                           REGION "RED OFF"
                               IF NOT "Clock_1Hz" THEN
                                   CASE #j OF
                                       #"Part 01":
                                           #stackLight := #stackLight AND (NOT #"Part 01 Red On");
                                           #stackLight := #stackLight AND (NOT #"Part 01 Yellow On");
                                           #stackLight := #stackLight AND (NOT #"Part 01 Green On");
                                       #"Part 02":
                                           #stackLight := #stackLight AND (NOT #"Part 02 Red On");
                                           #stackLight := #stackLight AND (NOT #"Part 02 Yellow On");
                                           #stackLight := #stackLight AND (NOT #"Part 02 Green On");
                                       #"Part 03":
                                           #stackLight := #stackLight AND (NOT #"Part 03 Red On");
                                           #stackLight := #stackLight AND (NOT #"Part 03 Yellow On");
                                           #stackLight := #stackLight AND (NOT #"Part 03 Green On");
                                       #"Part 04":
                                           #stackLight := #stackLight AND (NOT #"Part 04 Red On");
                                           #stackLight := #stackLight AND (NOT #"Part 04 Yellow On");
                                           #stackLight := #stackLight AND (NOT #"Part 04 Green On");
                                       #"Part 05":
                                           #stackLight := #stackLight AND (NOT #"Part 05 Red On");
                                           #stackLight := #stackLight AND (NOT #"Part 05 Yellow On");
                                           #stackLight := #stackLight AND (NOT #"Part 05 Green On");
                                       #"Part 06":
                                           #stackLight := #stackLight AND (NOT #"Part 06 Red On");
                                           #stackLight := #stackLight AND (NOT #"Part 06 Yellow On");
                                           #stackLight := #stackLight AND (NOT #"Part 06 Green On");
                                       ELSE
                                           ;
                                   END_CASE;
                               END_IF;
                           END_REGION

                       END_IF;
                   END_REGION

                   REGION "COPY OUT TO GLOBAL"
                       #stations.me[#i].stackLightOut := #stackLight;
                   END_REGION

               END_FOR;
           END_REGION

       END_FOR;
   END_REGION
END_FUNCTION_BLOCK

FUNCTION_BLOCK "KP8 Button Activation"   // FB12, SCL
{ S7_Optimized_Access := 'TRUE' }
VERSION : 0.1
   VAR_IN_OUT
      stations : "Stations";
   END_VAR
   VAR
      old : Struct
         kp8Config : Array[0.."stnCount"] of "KP8 Button Config";
      END_STRUCT;
   END_VAR
   VAR_TEMP
      btnCount : Int;
      currentPNs : Array[0..7] of WString[40];
      i : Int;
      init : Bool;
      j : Int;
      stnCount : Int;
      temp : Int;
   END_VAR
BEGIN
   REGION "GET STATION COUNT"
       #stnCount := "stnCount";
       #btnCount := "ptsPerStn";
   END_REGION

   REGION "LOOP THROUGH STATIONS"
       FOR #i := 0 TO #stnCount DO

           REGION "COPY TO LOCAL"
               #currentPNs := #stations.me[#i].partNumbers;
           END_REGION


           REGION "LOOP THROUGH BUTTONS"
               FOR #j := 0 TO #btnCount DO

                       REGION "ACTIVATE BUTTON"
                           IF LEN(#currentPNs[#j]) <> 0 THEN
                               #stations.me[#i].kp8Config.activate[#j] := TRUE;
                               #stations.me[#i].kp8Config.colorOff[#j] := 'green';
                               #stations.me[#i].kp8Config.colorOn1[#j] := 'yellow';
                               #stations.me[#i].kp8Config.colorOn2[#j] := '';
                               #stations.me[#i].kp8Config.flash[#j] := FALSE;
                               #stations.me[#i].kp8Config.group[#j] := 0;
                               #stations.me[#i].kp8Config.mode[#j] := TRUE;
                           END_IF;
                       END_REGION

                       REGION "DEACTIVATE BUTTON"
                           IF LEN(#currentPNs[#j]) = 0 THEN
                               #stations.me[#i].kp8Config.activate[#j] := FALSE;
                               #stations.me[#i].kp8Config.colorOff[#j] := '';
                               #stations.me[#i].kp8Config.colorOn1[#j] := '';
                               #stations.me[#i].kp8Config.colorOn2[#j] := '';
                               #stations.me[#i].kp8Config.flash[#j] := FALSE;
                               #stations.me[#i].kp8Config.group[#j] := 0;
                               #stations.me[#i].kp8Config.mode[#j] := FALSE;
                           END_IF;
                       END_REGION

               END_FOR;
           END_REGION

           REGION "SOFT INIT"
               IF #stations.me[#i].kp8Config <> #old.kp8Config[#i] THEN
                   #stations.me[#i].init.soft := TRUE;
               END_IF;
           END_REGION

           REGION "SAVE FOR CHANGE DETECTION"
               #old.kp8Config[#i] := #stations.me[#i].kp8Config;
           END_REGION

       END_FOR;
   END_REGION
END_FUNCTION_BLOCK

FUNCTION_BLOCK "Remove Part Request"   // FB13, SCL
{ S7_Optimized_Access := 'TRUE' }
VERSION : 0.1
   VAR_IN_OUT
      pRow : Int;
      requests : "Part Request Data";
      stations : "Stations";
   END_VAR
   VAR
      old : Struct
         partReq : "Station Old Presses";
      END_STRUCT;
   END_VAR
   VAR_TEMP
      address : UInt;
      blankRow : "Table Row";
      hasPart : Bool;
      i : Int;
      j : Int;
      k : Int;
      logAddress : UInt;
      maxRows : Int;
      noPart : Bool;
      oldPartReq : Bool;
      partNumber : WString;
      partReq : Bool;
      pRemoveRow : Int;
      btnCount : Int;
      stnCount : Int;
      removeAddress : Bool;
   END_VAR
BEGIN
   REGION "COPY TO LOCAL"
       #maxRows := "partReqHmiRowCount";
       #stnCount := "stnCount";
       #btnCount := "ptsPerStn";
   END_REGION


   REGION "FOR EACH STATION"
       FOR #i := 0 TO #stnCount DO

           REGION "FOR EACH BUTTON"
               FOR #j := 1 TO #btnCount DO

                   REGION "COPY TO LOCAL"
                       #partReq := #stations.me[#i].btnStates[#j];
                       #oldPartReq := #old.partReq.me[#i, #j];
                   END_REGION

                   REGION "DETERMINE STATE"

                       REGION "PART REQUEST FALLING EDGE"
                           IF NOT #partReq AND #oldPartReq THEN

                               REGION "SAVE FOR CHANGE DETECTION"
                                   #old.partReq.me[#i, #j] := #partReq;
                               END_REGION

                               REGION "COPY TO LOCAL"
                                   #partNumber := #stations.me[#i].partNumbers[#j];
                               END_REGION

                               REGION "BUTTON HAS NO PART"
                                   IF #partNumber = wstring#'' THEN
                                       #hasPart := FALSE;
                                       #noPart := TRUE;
                                   END_IF;
                               END_REGION

                               REGION "BUTTON HAS PART"
                                   IF #partNumber <> wstring#'' THEN
                                       #hasPart := TRUE;
                                       #noPart := FALSE;
                                   END_IF;
                               END_REGION

                           END_IF;
                       END_REGION

                   END_REGION

                   REGION "NO PART"
                       IF #noPart THEN

                           REGION "TURN OFF THE LIGHTS"
                               #hasPart := FALSE;
                               #noPart := FALSE;
                           END_REGION

                       END_IF;

                   END_REGION

                   REGION "HAS PART"
                       IF #hasPart THEN

                           REGION "TURN OFF THE LIGHTS"
                               #hasPart := FALSE;
                           END_REGION

                           REGION "CALCULATE ADDRESS"
                               #address := (INT_TO_UINT(#i) + 1) * 10 + (INT_TO_UINT(#j) + 1);
                           END_REGION

                           REGION "RESET FLAG"
                               #removeAddress := FALSE;
                           END_REGION

                           REGION "SEARCH EACH ROW IN PART DB"
                               FOR #k := 0 TO #maxRows DO

                                   REGION "COPY TO LOCAL"
                                       #logAddress := #requests.row[#k].address;
                                   END_REGION

                                   REGION "ON MATCH"
                                       IF #logAddress = #address THEN

                                           REGION "SET FLAG"
                                               #removeAddress := TRUE;
                                           END_REGION

                                           REGION "SAVE POINTER"
                                               #pRemoveRow := #k;
                                           END_REGION

                                       END_IF;
                                   END_REGION

                               END_FOR;
                           END_REGION

                       END_IF;
                   END_REGION

                   REGION "REMOVE ADDRESS"
                       IF #removeAddress THEN

                           REGION "TURN OFF THE LIGHTS"
                               #removeAddress := FALSE;
                           END_REGION

                           REGION "TURN OFF REQUEST"
                               #stations.me[#i].partRequested[#j] := FALSE;
                           END_REGION

                           REGION "REMOVAL PROCESS"

                               REGION "REMOVE ROW"
                                   #requests.row[#pRemoveRow] := #blankRow;
                               END_REGION

                               REGION "REMOVE PART ORDERED"
                                   #stations.me[#i].partOrdered[#j] := FALSE;
                               END_REGION

                           END_REGION

                           REGION "ROW POINTER"

                               REGION "DECREMENT"
                                   #pRow := #pRow - 1;
                               END_REGION

                               REGION "LOW LIMIT ROLL OVER"
                                   IF #pRow < 0 THEN
                                       #pRow := 0;
                                   END_IF;
                               END_REGION

                           END_REGION

                       END_IF;
                   END_REGION

               END_FOR;

           END_REGION

       END_FOR;
   END_REGION
END_FUNCTION_BLOCK

FUNCTION_BLOCK "HMI Settings Screen"   // FB14, LAD
{ S7_Optimized_Access := 'TRUE' }
VERSION : 0.1
   VAR_IN_OUT
      settings : "Settings";
      stations : "Stations";
   END_VAR
   VAR
      tmrTimeOut : TON_TIME;
      instStaSel : "Station Selection";
      instKP8BtnSel : "KP8 Button Selections";
      old : Struct
         asgnPN : Bool;
         asgnAlloted : Bool;
         asgnCritical : Bool;
         nextPress : Bool;
         prevPress : Bool;
         selBtnCount : Int;
         selBtnNumber : Int;
         selStnCount : Int;
         selStnNumber : Int;
      END_STRUCT;
      instAsnBtnPrms : "Assign Button Parameters";
      instAniPNTmr : "Animate: PN & Timers";
   END_VAR
   VAR_TEMP
      pBN : Int;
      pSN : Int;
      wStringBox : WString;
   END_VAR
   VAR CONSTANT
      ptTimeOut : Time := t#15m;
   END_VAR
   VAR_TEMP   // added for the SCL form of the ladder/FBD networks
      _w1 : Bool;
   END_VAR
BEGIN

REGION Network 1: ENTRY TIMEOUT
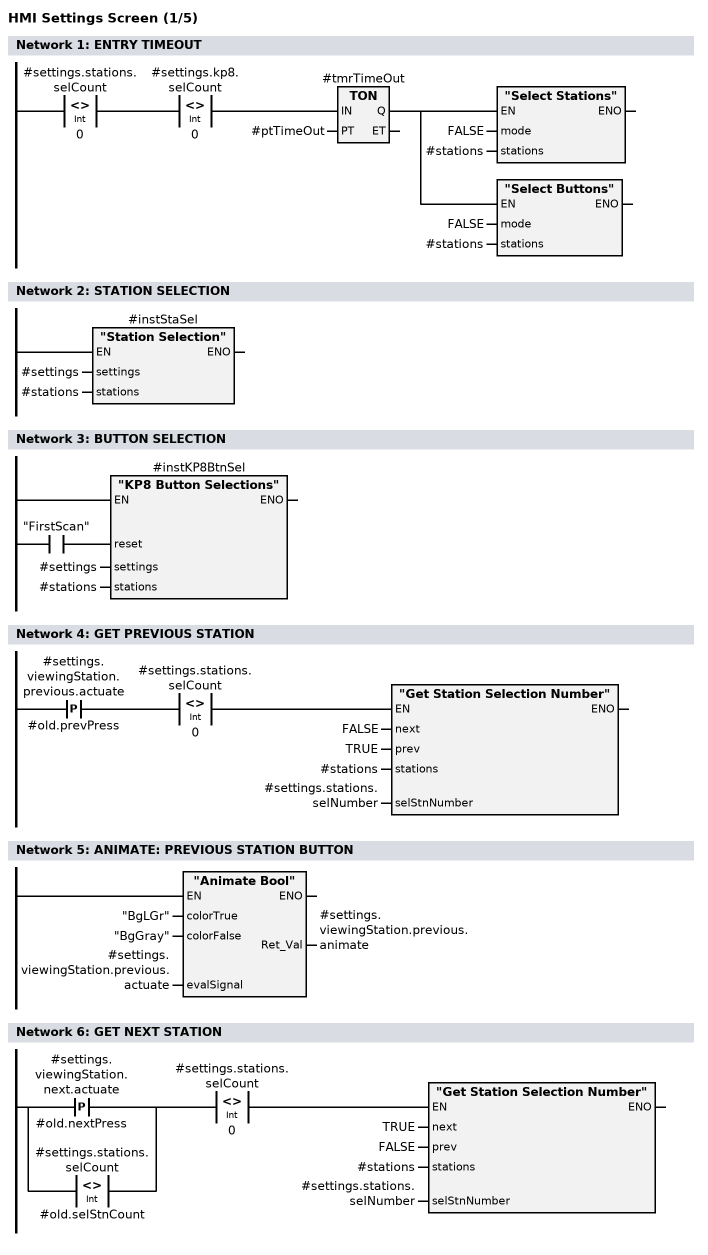
   #tmrTimeOut(IN := (#settings.stations.selCount <> 0) AND (#settings.kp8.selCount <> 0), PT := #ptTimeOut);   // TON
   IF #tmrTimeOut.Q THEN
       "Select Stations"(mode := FALSE, stations := #stations);
       "Select Buttons"(mode := FALSE, stations := #stations);
   END_IF;
END_REGION

REGION Network 2: STATION SELECTION
   RUNG wire#powerrail
      #instStaSel(settings := #settings, stations := #stations)
   END_RUNG
   // the same network as SCL:
   #instStaSel(settings := #settings, stations := #stations);   // "Station Selection"
END_REGION

REGION Network 3: BUTTON SELECTION
   RUNG wire#powerrail
      #instKP8BtnSel(reset := wire#w1, settings := #settings, stations := #stations)
   END_RUNG
   RUNG wire#powerrail
      Contact( "FirstScan" )
   END_RUNG wire#w1
   // the same network as SCL:
   #instKP8BtnSel(reset := "FirstScan", settings := #settings, stations := #stations);   // "KP8 Button Selections"
END_REGION

REGION Network 4: GET PREVIOUS STATION
   RUNG wire#powerrail
      P_Contact(operand := #settings.viewingStation.previous.actuate, bit := #old.prevPress)
      { S7_Templates := "SrcType := Int" } NE_Contact(in1 := #settings.stations.selCount, in2 := 0)
      "Get Station Selection Number"(next := FALSE, prev := TRUE, stations := #stations, selStnNumber := #settings.stations.selNumber)
   END_RUNG
   // the same network as SCL:
   #_w1 := #settings.viewingStation.previous.actuate AND NOT #old.prevPress;   // rising edge of #settings.viewingStation.previous.actuate
   #old.prevPress := #settings.viewingStation.previous.actuate;
   IF #_w1 AND (#settings.stations.selCount <> 0) THEN
       "Get Station Selection Number"(next := FALSE,
                               prev := TRUE,
                               stations := #stations,
                               selStnNumber := #settings.stations.selNumber);
   END_IF;
END_REGION

REGION Network 5: ANIMATE: PREVIOUS STATION BUTTON
   RUNG wire#powerrail
      "Animate Bool"(colorTrue := "BgLGr", colorFalse := "BgGray", evalSignal := #settings.viewingStation.previous.actuate, Ret_Val => #settings.viewingStation.previous.animate)
   END_RUNG
   // the same network as SCL:
   #settings.viewingStation.previous.animate := "Animate Bool"(colorTrue := "BgLGr",
                           colorFalse := "BgGray",
                           evalSignal := #settings.viewingStation.previous.actuate);
END_REGION

REGION Network 6: GET NEXT STATION
   RUNG wire#powerrail
      P_Contact(operand := #settings.viewingStation.next.actuate, bit := #old.nextPress)
      wire#w1
      { S7_Templates := "SrcType := Int" } NE_Contact(in1 := #settings.stations.selCount, in2 := 0)
      "Get Station Selection Number"(next := TRUE, prev := FALSE, stations := #stations, selStnNumber := #settings.stations.selNumber)
   END_RUNG
   RUNG wire#powerrail
      { S7_Templates := "SrcType := Int" } NE_Contact(in1 := #settings.stations.selCount, in2 := #old.selStnCount)
   END_RUNG wire#w1
   // the same network as SCL:
   #_w1 := #settings.viewingStation.next.actuate AND NOT #old.nextPress;   // rising edge of #settings.viewingStation.next.actuate
   #old.nextPress := #settings.viewingStation.next.actuate;
   IF (#_w1 OR (#settings.stations.selCount <> #old.selStnCount)) AND (#settings.stations.selCount <> 0) THEN
       "Get Station Selection Number"(next := TRUE,
                               prev := FALSE,
                               stations := #stations,
                               selStnNumber := #settings.stations.selNumber);
   END_IF;
END_REGION

REGION Network 7: ANIMATE: NEXT STATION BUTTON
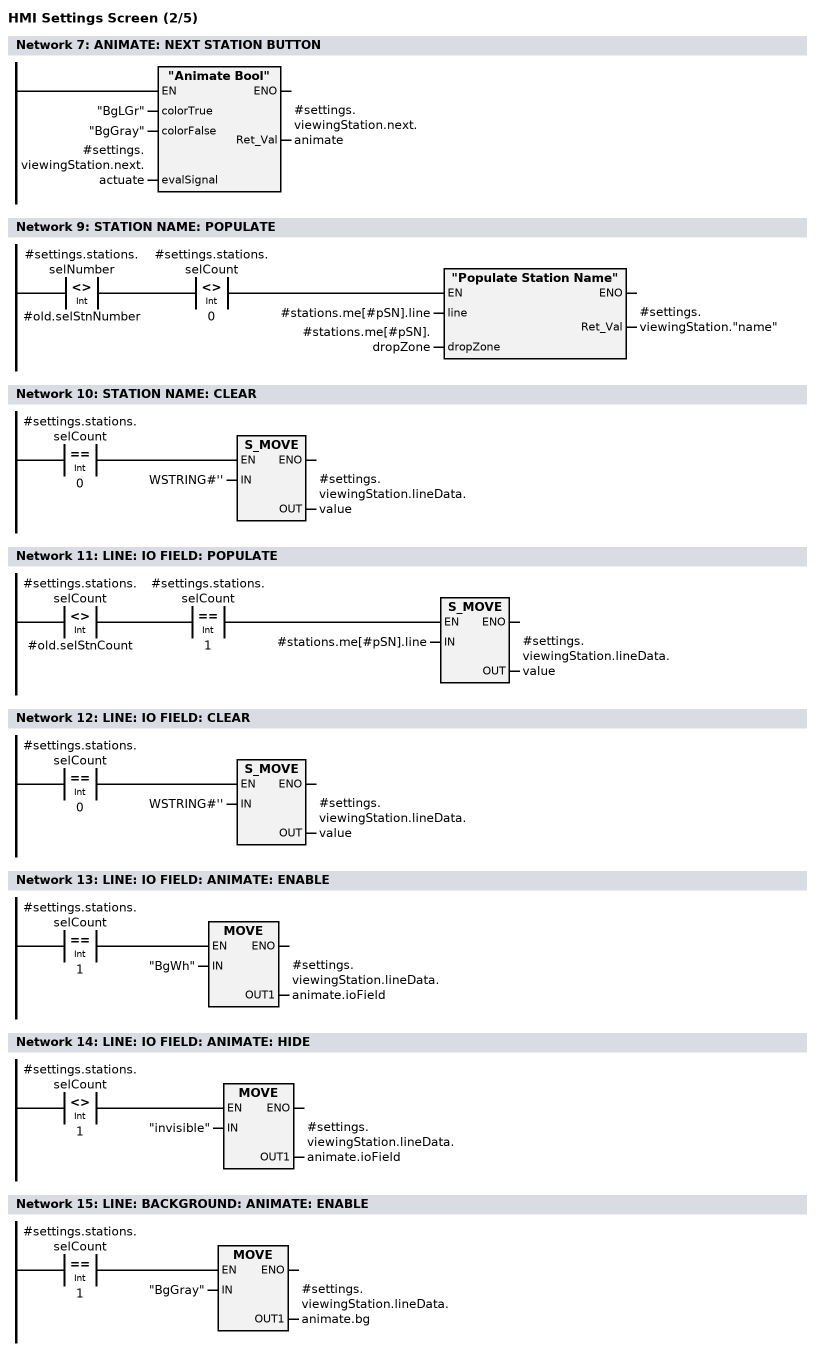
   RUNG wire#powerrail
      "Animate Bool"(colorTrue := "BgLGr", colorFalse := "BgGray", evalSignal := #settings.viewingStation.next.actuate, Ret_Val => #settings.viewingStation.next.animate)
   END_RUNG
   // the same network as SCL:
   #settings.viewingStation.next.animate := "Animate Bool"(colorTrue := "BgLGr",
                           colorFalse := "BgGray",
                           evalSignal := #settings.viewingStation.next.actuate);
END_REGION

REGION Network 8 (SCL): COPY TO POINTERS
   #pSN := #settings.stations.selNumber;
   #pBN := #settings.kp8.selBtnNumber;
END_REGION

REGION Network 9: STATION NAME: POPULATE
   RUNG wire#powerrail
      { S7_Templates := "SrcType := Int" } NE_Contact(in1 := #settings.stations.selNumber, in2 := #old.selStnNumber)
      { S7_Templates := "SrcType := Int" } NE_Contact(in1 := #settings.stations.selCount, in2 := 0)
      "Populate Station Name"(line := #stations.me[#pSN].line, dropZone := #stations.me[#pSN].dropZone, Ret_Val => #settings.viewingStation."name")
   END_RUNG
   // the same network as SCL:
   IF (#settings.stations.selNumber <> #old.selStnNumber) AND (#settings.stations.selCount <> 0) THEN
       #settings.viewingStation."name" := "Populate Station Name"(line := #stations.me[#pSN].line,
                               dropZone := #stations.me[#pSN].dropZone);
   END_IF;
END_REGION

REGION Network 10: STATION NAME: CLEAR
   RUNG wire#powerrail
      { S7_Templates := "SrcType := Int" } EQ_Contact(in1 := #settings.stations.selCount, in2 := 0)
      S_Move(in := WSTRING#'', out => #settings.viewingStation.lineData.value)
   END_RUNG
   // the same network as SCL:
   IF #settings.stations.selCount = 0 THEN #settings.viewingStation.lineData.value := WSTRING#''; END_IF;
END_REGION

REGION Network 11: LINE: IO FIELD: POPULATE
   RUNG wire#powerrail
      { S7_Templates := "SrcType := Int" } NE_Contact(in1 := #settings.stations.selCount, in2 := #old.selStnCount)
      { S7_Templates := "SrcType := Int" } EQ_Contact(in1 := #settings.stations.selCount, in2 := 1)
      S_Move(in := #stations.me[#pSN].line, out => #settings.viewingStation.lineData.value)
   END_RUNG
   // the same network as SCL:
   IF (#settings.stations.selCount <> #old.selStnCount) AND (#settings.stations.selCount = 1) THEN
       #settings.viewingStation.lineData.value := #stations.me[#pSN].line;
   END_IF;
END_REGION

REGION Network 12: LINE: IO FIELD: CLEAR
   RUNG wire#powerrail
      { S7_Templates := "SrcType := Int" } EQ_Contact(in1 := #settings.stations.selCount, in2 := 0)
      S_Move(in := WSTRING#'', out => #settings.viewingStation.lineData.value)
   END_RUNG
   // the same network as SCL:
   IF #settings.stations.selCount = 0 THEN #settings.viewingStation.lineData.value := WSTRING#''; END_IF;
END_REGION

REGION Network 13: LINE: IO FIELD: ANIMATE: ENABLE
   RUNG wire#powerrail
      { S7_Templates := "SrcType := Int" } EQ_Contact(in1 := #settings.stations.selCount, in2 := 1)
      Move(in := "BgWh", out1 => #settings.viewingStation.lineData.animate.ioField)
   END_RUNG
   // the same network as SCL:
   IF #settings.stations.selCount = 1 THEN
       #settings.viewingStation.lineData.animate.ioField := "BgWh";
   END_IF;
END_REGION

REGION Network 14: LINE: IO FIELD: ANIMATE: HIDE
   RUNG wire#powerrail
      { S7_Templates := "SrcType := Int" } NE_Contact(in1 := #settings.stations.selCount, in2 := 1)
      Move(in := "invisible", out1 => #settings.viewingStation.lineData.animate.ioField)
   END_RUNG
   // the same network as SCL:
   IF #settings.stations.selCount <> 1 THEN
       #settings.viewingStation.lineData.animate.ioField := "invisible";
   END_IF;
END_REGION

REGION Network 15: LINE: BACKGROUND: ANIMATE: ENABLE
   RUNG wire#powerrail
      { S7_Templates := "SrcType := Int" } EQ_Contact(in1 := #settings.stations.selCount, in2 := 1)
      Move(in := "BgGray", out1 => #settings.viewingStation.lineData.animate.bg)
   END_RUNG
   // the same network as SCL:
   IF #settings.stations.selCount = 1 THEN #settings.viewingStation.lineData.animate.bg := "BgGray"; END_IF;
END_REGION

REGION Network 16: LINE: BACKGROUND: ANIMATE: HIDE
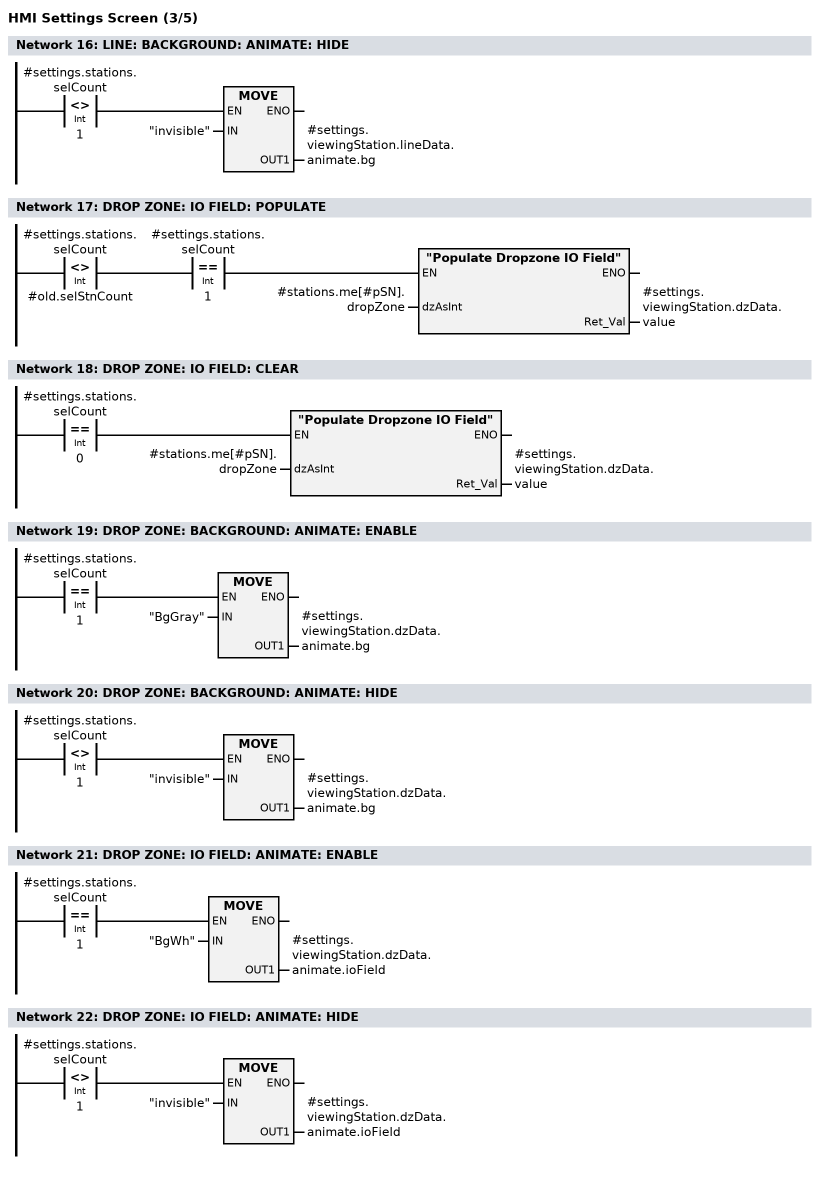
   RUNG wire#powerrail
      { S7_Templates := "SrcType := Int" } NE_Contact(in1 := #settings.stations.selCount, in2 := 1)
      Move(in := "invisible", out1 => #settings.viewingStation.lineData.animate.bg)
   END_RUNG
   // the same network as SCL:
   IF #settings.stations.selCount <> 1 THEN
       #settings.viewingStation.lineData.animate.bg := "invisible";
   END_IF;
END_REGION

REGION Network 17: DROP ZONE: IO FIELD: POPULATE
   RUNG wire#powerrail
      { S7_Templates := "SrcType := Int" } NE_Contact(in1 := #settings.stations.selCount, in2 := #old.selStnCount)
      { S7_Templates := "SrcType := Int" } EQ_Contact(in1 := #settings.stations.selCount, in2 := 1)
      "Populate Dropzone IO Field"(dzAsInt := #stations.me[#pSN].dropZone, Ret_Val => #settings.viewingStation.dzData.value)
   END_RUNG
   // the same network as SCL:
   IF (#settings.stations.selCount <> #old.selStnCount) AND (#settings.stations.selCount = 1) THEN
       #settings.viewingStation.dzData.value := "Populate Dropzone IO Field"(dzAsInt := #stations.me[#pSN].dropZone);
   END_IF;
END_REGION

REGION Network 18: DROP ZONE: IO FIELD: CLEAR
   RUNG wire#powerrail
      { S7_Templates := "SrcType := Int" } EQ_Contact(in1 := #settings.stations.selCount, in2 := 0)
      "Populate Dropzone IO Field"(dzAsInt := #stations.me[#pSN].dropZone, Ret_Val => #settings.viewingStation.dzData.value)
   END_RUNG
   // the same network as SCL:
   IF #settings.stations.selCount = 0 THEN
       #settings.viewingStation.dzData.value := "Populate Dropzone IO Field"(dzAsInt := #stations.me[#pSN].dropZone);
   END_IF;
END_REGION

REGION Network 19: DROP ZONE: BACKGROUND: ANIMATE: ENABLE
   RUNG wire#powerrail
      { S7_Templates := "SrcType := Int" } EQ_Contact(in1 := #settings.stations.selCount, in2 := 1)
      Move(in := "BgGray", out1 => #settings.viewingStation.dzData.animate.bg)
   END_RUNG
   // the same network as SCL:
   IF #settings.stations.selCount = 1 THEN #settings.viewingStation.dzData.animate.bg := "BgGray"; END_IF;
END_REGION

REGION Network 20: DROP ZONE: BACKGROUND: ANIMATE: HIDE
   RUNG wire#powerrail
      { S7_Templates := "SrcType := Int" } NE_Contact(in1 := #settings.stations.selCount, in2 := 1)
      Move(in := "invisible", out1 => #settings.viewingStation.dzData.animate.bg)
   END_RUNG
   // the same network as SCL:
   IF #settings.stations.selCount <> 1 THEN
       #settings.viewingStation.dzData.animate.bg := "invisible";
   END_IF;
END_REGION

REGION Network 21: DROP ZONE: IO FIELD: ANIMATE: ENABLE
   RUNG wire#powerrail
      { S7_Templates := "SrcType := Int" } EQ_Contact(in1 := #settings.stations.selCount, in2 := 1)
      Move(in := "BgWh", out1 => #settings.viewingStation.dzData.animate.ioField)
   END_RUNG
   // the same network as SCL:
   IF #settings.stations.selCount = 1 THEN #settings.viewingStation.dzData.animate.ioField := "BgWh"; END_IF;
END_REGION

REGION Network 22: DROP ZONE: IO FIELD: ANIMATE: HIDE
   RUNG wire#powerrail
      { S7_Templates := "SrcType := Int" } NE_Contact(in1 := #settings.stations.selCount, in2 := 1)
      Move(in := "invisible", out1 => #settings.viewingStation.dzData.animate.ioField)
   END_RUNG
   // the same network as SCL:
   IF #settings.stations.selCount <> 1 THEN
       #settings.viewingStation.dzData.animate.ioField := "invisible";
   END_IF;
END_REGION

REGION Network 23: PART NUMBER IO FIELD: POPULATE
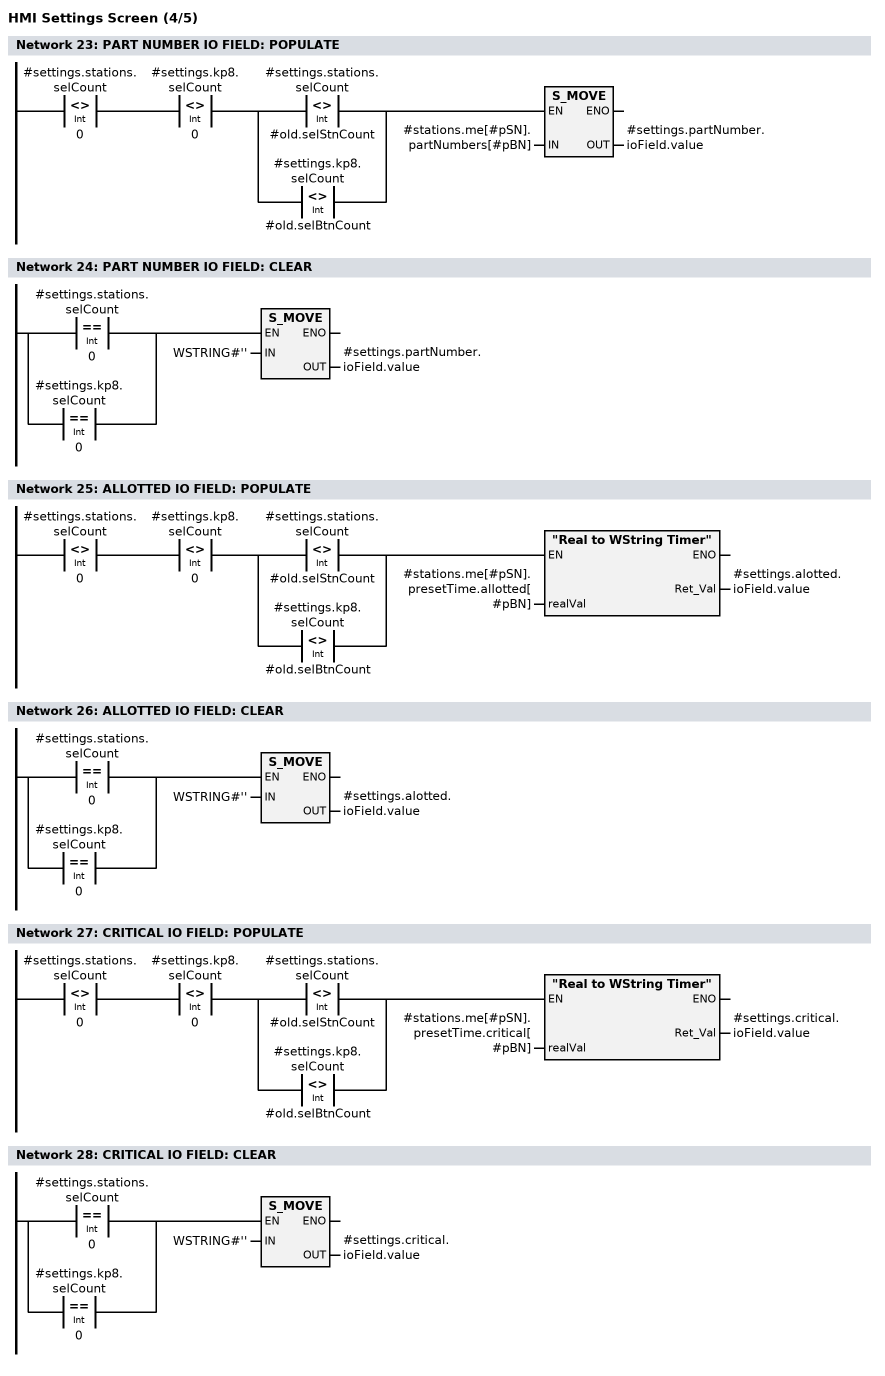
   RUNG wire#powerrail
      { S7_Templates := "SrcType := Int" } NE_Contact(in1 := #settings.stations.selCount, in2 := 0)
      { S7_Templates := "SrcType := Int" } NE_Contact(in1 := #settings.kp8.selCount, in2 := 0)
      wire#w1
      { S7_Templates := "SrcType := Int" } NE_Contact(in1 := #settings.stations.selCount, in2 := #old.selStnCount)
      wire#w2
      S_Move(in := #stations.me[#pSN].partNumbers[#pBN], out => #settings.partNumber.ioField.value)
   END_RUNG
   RUNG wire#w1
      { S7_Templates := "SrcType := Int" } NE_Contact(in1 := #settings.kp8.selCount, in2 := #old.selBtnCount)
   END_RUNG wire#w2
   // the same network as SCL:
   IF (#settings.stations.selCount <> 0) AND (#settings.kp8.selCount <> 0) AND ((#settings.stations.selCount <> #old.selStnCount) OR (#settings.kp8.selCount <> #old.selBtnCount)) THEN
       #settings.partNumber.ioField.value := #stations.me[#pSN].partNumbers[#pBN];
   END_IF;
END_REGION

REGION Network 24: PART NUMBER IO FIELD: CLEAR
   RUNG wire#powerrail
      { S7_Templates := "SrcType := Int" } EQ_Contact(in1 := #settings.stations.selCount, in2 := 0)
      wire#w1
      S_Move(in := WSTRING#'', out => #settings.partNumber.ioField.value)
   END_RUNG
   RUNG wire#powerrail
      { S7_Templates := "SrcType := Int" } EQ_Contact(in1 := #settings.kp8.selCount, in2 := 0)
   END_RUNG wire#w1
   // the same network as SCL:
   IF (#settings.stations.selCount = 0) OR (#settings.kp8.selCount = 0) THEN
       #settings.partNumber.ioField.value := WSTRING#'';
   END_IF;
END_REGION

REGION Network 25: ALLOTTED IO FIELD: POPULATE
   RUNG wire#powerrail
      { S7_Templates := "SrcType := Int" } NE_Contact(in1 := #settings.stations.selCount, in2 := 0)
      { S7_Templates := "SrcType := Int" } NE_Contact(in1 := #settings.kp8.selCount, in2 := 0)
      wire#w1
      { S7_Templates := "SrcType := Int" } NE_Contact(in1 := #settings.stations.selCount, in2 := #old.selStnCount)
      wire#w2
      "Real to WString Timer"(realVal := #stations.me[#pSN].presetTime.allotted[#pBN], Ret_Val => #settings.alotted.ioField.value)
   END_RUNG
   RUNG wire#w1
      { S7_Templates := "SrcType := Int" } NE_Contact(in1 := #settings.kp8.selCount, in2 := #old.selBtnCount)
   END_RUNG wire#w2
   // the same network as SCL:
   IF (#settings.stations.selCount <> 0) AND (#settings.kp8.selCount <> 0) AND ((#settings.stations.selCount <> #old.selStnCount) OR (#settings.kp8.selCount <> #old.selBtnCount)) THEN
       #settings.alotted.ioField.value := "Real to WString Timer"(realVal := #stations.me[#pSN].presetTime.allotted[#pBN]);
   END_IF;
END_REGION

REGION Network 26: ALLOTTED IO FIELD: CLEAR
   RUNG wire#powerrail
      { S7_Templates := "SrcType := Int" } EQ_Contact(in1 := #settings.stations.selCount, in2 := 0)
      wire#w1
      S_Move(in := WSTRING#'', out => #settings.alotted.ioField.value)
   END_RUNG
   RUNG wire#powerrail
      { S7_Templates := "SrcType := Int" } EQ_Contact(in1 := #settings.kp8.selCount, in2 := 0)
   END_RUNG wire#w1
   // the same network as SCL:
   IF (#settings.stations.selCount = 0) OR (#settings.kp8.selCount = 0) THEN
       #settings.alotted.ioField.value := WSTRING#'';
   END_IF;
END_REGION

REGION Network 27: CRITICAL IO FIELD: POPULATE
   RUNG wire#powerrail
      { S7_Templates := "SrcType := Int" } NE_Contact(in1 := #settings.stations.selCount, in2 := 0)
      { S7_Templates := "SrcType := Int" } NE_Contact(in1 := #settings.kp8.selCount, in2 := 0)
      wire#w1
      { S7_Templates := "SrcType := Int" } NE_Contact(in1 := #settings.stations.selCount, in2 := #old.selStnCount)
      wire#w2
      "Real to WString Timer"(realVal := #stations.me[#pSN].presetTime.critical[#pBN], Ret_Val => #settings.critical.ioField.value)
   END_RUNG
   RUNG wire#w1
      { S7_Templates := "SrcType := Int" } NE_Contact(in1 := #settings.kp8.selCount, in2 := #old.selBtnCount)
   END_RUNG wire#w2
   // the same network as SCL:
   IF (#settings.stations.selCount <> 0) AND (#settings.kp8.selCount <> 0) AND ((#settings.stations.selCount <> #old.selStnCount) OR (#settings.kp8.selCount <> #old.selBtnCount)) THEN
       #settings.critical.ioField.value := "Real to WString Timer"(realVal := #stations.me[#pSN].presetTime.critical[#pBN]);
   END_IF;
END_REGION

REGION Network 28: CRITICAL IO FIELD: CLEAR
   RUNG wire#powerrail
      { S7_Templates := "SrcType := Int" } EQ_Contact(in1 := #settings.stations.selCount, in2 := 0)
      wire#w1
      S_Move(in := WSTRING#'', out => #settings.critical.ioField.value)
   END_RUNG
   RUNG wire#powerrail
      { S7_Templates := "SrcType := Int" } EQ_Contact(in1 := #settings.kp8.selCount, in2 := 0)
   END_RUNG wire#w1
   // the same network as SCL:
   IF (#settings.stations.selCount = 0) OR (#settings.kp8.selCount = 0) THEN
       #settings.critical.ioField.value := WSTRING#'';
   END_IF;
END_REGION

REGION Network 29: PART NUMBER, ALLOTTED & CRITICAL: ANIMATE
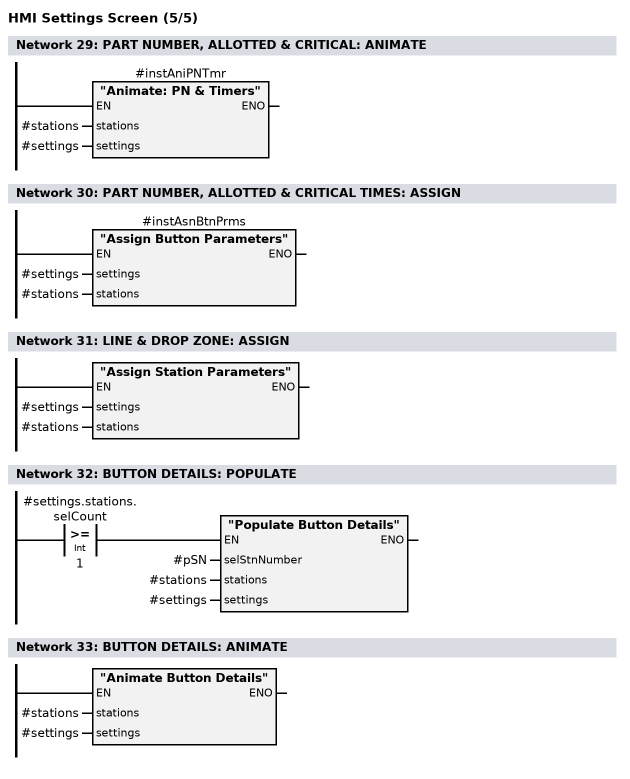
   RUNG wire#powerrail
      #instAniPNTmr(stations := #stations, settings := #settings)
   END_RUNG
   // the same network as SCL:
   #instAniPNTmr(stations := #stations, settings := #settings);   // "Animate: PN & Timers"
END_REGION

REGION Network 30: PART NUMBER, ALLOTTED & CRITICAL TIMES: ASSIGN
   RUNG wire#powerrail
      #instAsnBtnPrms(settings := #settings, stations := #stations)
   END_RUNG
   // the same network as SCL:
   #instAsnBtnPrms(settings := #settings, stations := #stations);   // "Assign Button Parameters"
END_REGION

REGION Network 31: LINE & DROP ZONE: ASSIGN
   RUNG wire#powerrail
      "Assign Station Parameters"(settings := #settings, stations := #stations)
   END_RUNG
   // the same network as SCL:
   "Assign Station Parameters"(settings := #settings, stations := #stations);
END_REGION

REGION Network 32: BUTTON DETAILS: POPULATE
   RUNG wire#powerrail
      { S7_Templates := "SrcType := Int" } GE_Contact(in1 := #settings.stations.selCount, in2 := 1)
      "Populate Button Details"(selStnNumber := #pSN, stations := #stations, settings := #settings)
   END_RUNG
   // the same network as SCL:
   IF #settings.stations.selCount >= 1 THEN
       "Populate Button Details"(selStnNumber := #pSN, stations := #stations, settings := #settings);
   END_IF;
END_REGION

REGION Network 33: BUTTON DETAILS: ANIMATE
   RUNG wire#powerrail
      "Animate Button Details"(stations := #stations, settings := #settings)
   END_RUNG
   // the same network as SCL:
   "Animate Button Details"(stations := #stations, settings := #settings);
END_REGION

REGION Network 34 (SCL): CHANGE DETECTION
   #old.selBtnCount := #settings.kp8.selCount;
   #old.selBtnNumber := #settings.kp8.selBtnNumber;
   #old.selStnCount := #settings.stations.selCount;
   #old.selStnNumber := #settings.stations.selNumber;
END_REGION
END_FUNCTION_BLOCK

FUNCTION_BLOCK "Collapse Table"   // FB15, SCL
{ S7_Optimized_Access := 'TRUE' }
VERSION : 0.1
   VAR_IN_OUT
      requests : "Part Request Data";
   END_VAR
   VAR
      tableBox : "Part Request Data";
   END_VAR
   VAR_TEMP
      address : Int;
      blankRow : "Table Row";
      collapseReq : Bool;
      i : Int;
      maxRows : Int;
      pCollapse : Int;
   END_VAR
BEGIN
   REGION "COPY TO LOCAL"
       #maxRows := "partReqHmiRowCount";
   END_REGION

   REGION "REMOVE EMPTY ROWS"

       REGION "FOR EACH ROW IN PART DB"
           FOR #i := 0 TO #maxRows DO

               REGION "COPY TO LOCAL"
                   #address := UINT_TO_INT(#requests.row[#i].address);
               END_REGION

               REGION "ROW IS NOT EMPTY"
                   IF #address <> 0 THEN

                       REGION "MOVE TO TEMP TABLE"
                           #tableBox.row[#pCollapse] := #requests.row[#i];
                       END_REGION

                       REGION "CALCULATE POINTER"
                           #pCollapse += 1;
                       END_REGION

                   END_IF;
               END_REGION

               REGION "ROW IS EMPTY"
                   IF #address = 0 THEN

                       REGION "SET FLAG"
                           #collapseReq := TRUE;
                       END_REGION

                   END_IF;
               END_REGION

           END_FOR;
       END_REGION

   END_REGION

   REGION "COLLAPSE TABLE"
       IF #collapseReq THEN

           REGION "TURN OFF THE LIGHTS"
               #collapseReq := FALSE;
           END_REGION

           REGION "COPY TEMP TO PERMANENT"
               #requests := #tableBox;
           END_REGION

           REGION "CLEAR VALUES FROM TEMP TABLE"
               FOR #i := 0 TO #maxRows DO
                   #tableBox.row[#i] := #blankRow;
               END_FOR;
           END_REGION
       END_IF;

   END_REGION
END_FUNCTION_BLOCK

FUNCTION_BLOCK "HMI Populate Part Call"   // FB16, SCL
{ S7_Optimized_Access := 'TRUE' }
VERSION : 0.1
   VAR_INPUT
      currentRowCount : Int;
      requests : "Part Request Data";
   END_VAR
   VAR_IN_OUT
      partCall : "Part Call Screen";
      tableNav : "Table Nav";
   END_VAR
   VAR
      firstRow : Int;
      old : Struct
         top : Bool;
         pgUp : Bool;
         lnUp : Bool;
         lnDn : Bool;
         pgDn : Bool;
         btm : Bool;
      END_STRUCT;
   END_VAR
   VAR_TEMP
      animate : Bool;
      btn : Struct
         top : Bool;
         pgUp : Bool;
         lnUp : Bool;
         lnDn : Bool;
         pgDn : Bool;
         btm : Bool;
      END_STRUCT;
      gray : USInt;
      green : USInt;
      i : Int;
      maxDBRows : Int;
      pRow : Int;
      visibleRows : Int;
      thisRow : Int;
      saveAct : Bool;
   END_VAR
BEGIN
   REGION "COPY TO LOCAL"
       #visibleRows := "partReqHmiRowCount";
       #maxDBRows := #currentRowCount;
       #btn.top := #tableNav.top.actuate;
       #btn.pgUp := #tableNav.pageUp.actuate;
       #btn.lnUp := #tableNav.lineUp.actuate;
       #btn.lnDn := #tableNav.lineDown.actuate;
       #btn.pgDn := #tableNav.pageDown.actuate;
       #btn.btm := #tableNav.bottom.actuate;
   END_REGION

   REGION "RESOLVE FIRST ROW"

       REGION "TOP"
           IF NOT #btn.top AND #old.top THEN
               #firstRow := 0;
           END_IF;
       END_REGION

       REGION "PAGE UP"
           IF NOT #btn.pgUp AND #old.pgUp THEN
               #firstRow -= #visibleRows - 1;
           END_IF;
       END_REGION

       REGION "LINE UP"
           IF NOT #btn.lnUp AND #old.lnUp THEN
               #firstRow -= 1;
           END_IF;
       END_REGION

       REGION "LINE DOWN"
           IF NOT #btn.lnDn AND #old.lnDn THEN
               #firstRow += 1;
           END_IF;
       END_REGION

       REGION "PAGE DOWN"
           IF NOT #btn.pgDn AND #old.pgDn THEN
               #firstRow += #visibleRows - 1;
           END_IF;
       END_REGION

       REGION "BOTTOM"
           IF NOT #btn.btm AND #old.btm THEN
               #firstRow := #maxDBRows - #visibleRows + 1;
           END_IF;
       END_REGION

   END_REGION

   REGION "CHANGE DETECTION"
       #old.top := #btn.top;
       #old.pgUp := #btn.pgUp;
       #old.lnUp := #btn.lnUp;
       #old.lnDn := #btn.lnDn;
       #old.pgDn := #btn.pgDn;
       #old.btm := #btn.btm;
   END_REGION

   REGION "ANIMATE PART CALL NAV"

       REGION "COPY TO LOCAL"
           #gray := "BgGray";
           #green := "BgLGr";
       END_REGION

       REGION "TOP"
           #tableNav.top.animate := "Animate Bool"(colorTrue := #green,
                                                   colorFalse := #gray,
                                                   evalSignal := #tableNav.top.actuate);
       END_REGION

       REGION "PAGE UP"
           #tableNav.pageUp.animate := "Animate Bool"(colorTrue := #green,
                                                      colorFalse := #gray,
                                                      evalSignal := #tableNav.pageUp.actuate);
       END_REGION

       REGION "LINE UP"
           #tableNav.lineUp.animate := "Animate Bool"(colorTrue := #green,
                                                      colorFalse := #gray,
                                                      evalSignal := #tableNav.lineUp.actuate);
       END_REGION

       REGION "LINE DOWN"
           #tableNav.lineDown.animate := "Animate Bool"(colorTrue := #green,
                                                        colorFalse := #gray,
                                                        evalSignal := #tableNav.lineDown.actuate);
       END_REGION

       REGION "PAGE DOWN"
           #tableNav.pageDown.animate := "Animate Bool"(colorTrue := #green,
                                                        colorFalse := #gray,
                                                        evalSignal := #tableNav.pageDown.actuate);
       END_REGION

       REGION "BOTTOM"
           #tableNav.bottom.animate := "Animate Bool"(colorTrue := #green,
                                                      colorFalse := #gray,
                                                      evalSignal := #tableNav.bottom.actuate);
       END_REGION

   END_REGION

   REGION "UPPER LIMIT ROLL OVER"
       IF #firstRow > #maxDBRows THEN
           #firstRow -= #maxDBRows - 1;
       END_IF;
   END_REGION

   REGION "LOWER LIMIT ROLL OVER"
       IF #firstRow < 0 THEN
           #firstRow += #maxDBRows - 1;
       END_IF;
   END_REGION

   REGION "LOOP THROUGH DISPLAYED STATIONS"
       FOR #i := 0 TO #visibleRows - 1 DO

           REGION "CALCULATE POINTER"
               #pRow := #firstRow + #i;
           END_REGION

           REGION "UPPER LIMIT ROLL OVER"
               IF #maxDBRows <= #visibleRows THEN
                   #pRow := #i;
               END_IF;
               IF #pRow >= #maxDBRows AND #maxDBRows >= #visibleRows THEN
                   #pRow := #firstRow + #i - #maxDBRows;
               END_IF;
           END_REGION

           REGION "SEND TO HMI"
               #saveAct := #partCall.row[#i].pbSelection.actuate;
               #partCall.row[#i] := #requests.row[#pRow];
               #partCall.row[#i].pbSelection.actuate := #saveAct;
           END_REGION

       END_FOR;
   END_REGION
END_FUNCTION_BLOCK

FUNCTION_BLOCK "Clear Part Requests"   // FB17, SCL
{ S7_Optimized_Access := 'TRUE' }
VERSION : 0.1
   VAR_INPUT
      clearRequest : Bool;
   END_VAR
   VAR_IN_OUT
      requests : "Part Request Data";
      partCall : "Part Call Screen";
      currentRowCount : Int;
   END_VAR
   VAR_TEMP
      blankRow : "Table Row";
      i : Int;
      maxRows : Int;
   END_VAR
BEGIN
   REGION "ON REQUEST"
       IF #clearRequest THEN

           REGION "HMI TABLE"

               REGION "COPY TO LOCAL"
                   #maxRows := "partReqHmiRowCount";
               END_REGION

               REGION "CLEAR ROWS"
                   FOR #i := 0 TO #maxRows DO
                       #partCall.row[#i] := #blankRow;
                   END_FOR;
               END_REGION

           END_REGION

           REGION "PART REQUEST DATA BASE"

               REGION "COPY TO LOCAL"
                   #maxRows := "partReqDataRowCount";
               END_REGION

               REGION "CLEAR ROWS"
                   FOR #i := 0 TO #maxRows DO
                       #requests.row[#i] := #blankRow;
                       #currentRowCount := 0;
                   END_FOR;
               END_REGION

           END_REGION

       END_IF;
   END_REGION
END_FUNCTION_BLOCK

FUNCTION_BLOCK "Load Default Timer Presets"   // FB18, SCL
{ S7_Optimized_Access := 'TRUE' }
VERSION : 0.1
   VAR_INPUT
      req : Bool;
   END_VAR
   VAR_IN_OUT
      stations : "Stations";
   END_VAR
   VAR
      oldReq : Bool;
   END_VAR
   VAR_TEMP
      alotted : Real;
      btnCount : Int;
      critical : Real;
      i : Int;
      j : Int;
      partNumber : WString;
      stnCount : Int;
      tmrReal : Real;
   END_VAR
BEGIN
   REGION "COPY TO LOCAL"
       #alotted := "defaultAlotted";
       #btnCount := "ptsPerStn";
       #critical := "defaultCritical";
       #stnCount := #stnCount;
   END_REGION

   REGION "ON REQUEST RISING EDGE"
       IF #req AND NOT #oldReq THEN

           REGION "LOOP THROUGH STATIONS" 
               FOR #i := 0 TO #stnCount DO

                   REGION "LOOP THROUGH BUTTONS"
                       FOR #j := 0 TO #btnCount DO

                           REGION "COPY TO LOCAL"
                               #partNumber := #stations.me[#i].partNumbers[#j];
                           END_REGION

                           REGION "IF BUTTON HAS ASSOCIATED PN"
                               IF LEN(#partNumber) <> 0 THEN

                                   REGION "COPY TO LOCAL"
                                       #tmrReal := #stations.me[#i].presetTime.allotted[#j];
                                   END_REGION

                                   REGION "ON NO TIME ENTERED"
                                       IF #tmrReal = 0.0 THEN

                                           REGION "ASSIGN ALLOTTED VALUES"
                                               #stations.me[#i].presetTime.allotted[#j] := #alotted;
                                           END_REGION

                                       END_IF;
                                   END_REGION

                                   REGION "COPY TO LOCAL"
                                       #tmrReal := #stations.me[#i].presetTime.critical[#j];
                                   END_REGION

                                   REGION "ON NO TIME ENTERED"
                                       IF #tmrReal = 0.0 THEN

                                           REGION "ASSIGN CRITICAL VALUES"
                                               #stations.me[#i].presetTime.critical[#j] := #critical;
                                           END_REGION

                                       END_IF;
                                   END_REGION

                               END_IF;
                           END_REGION

                       END_FOR;
                   END_REGION

               END_FOR;
           END_REGION

       END_IF;
   END_REGION

   REGION "CHANGE DETECTION"
       #oldReq := #req;
   END_REGION ;
END_FUNCTION_BLOCK

FUNCTION_BLOCK "LED Populate Sign"   // FB19, SCL
{ S7_Optimized_Access := 'TRUE' }
VERSION : 0.1
   VAR_INPUT
      requests : "Part Request Data";
   END_VAR
   VAR_IN_OUT
      ledData : "LED Sign Data";
   END_VAR
   VAR_TEMP
      animate : USInt;
      i : Int;
      visibleRows : Int;
      tempRow : "Table Row";
   END_VAR
BEGIN
   REGION "COPY TO LOCAL"
       #visibleRows := "ledRowCount";
   END_REGION

   REGION "POPULATE SIGN DATA"

       REGION "FOR EACH ROW ON SIGN"
           FOR #i := 0 TO #visibleRows DO

               REGION "GET ROW"
                   #tempRow := #requests.row[#i];
               END_REGION

               REGION "LINE LABEL DARK MODE"                
                   "Dark Mode"(#tempRow.tfLine.animate);
               END_REGION